// TIA Portal project "CHM_BORDEIRA_20190721" (V15) (continued)
REGION Network 14: I1.5 - CSW Valve Closed (CV-311)
   // True = CLOSED, False = NOT
   RUNG wire#powerrail
      Contact( "CSW Valve Closed" )
      I_Contact( "CSW Valve Open" )
      Coil( "10_DI_Data".CV311_CLSD )
   END_RUNG
   // the same network as SCL:
   "10_DI_Data".CV311_CLSD := "CSW Valve Closed" AND NOT "CSW Valve Open";
END_REGION

REGION Network 15: I1.6 - Flue Gas Scrubber CSW Valve Open (CV-312)
   // True = OPEN, False = NOT
   RUNG wire#powerrail
      Contact( "Flue Gas Scrubber CSW Valve Opened" )
      I_Contact( "Flue Gas Scrubber CSW Valve Closed" )
      Coil( "10_DI_Data".CV312_OPN )
   END_RUNG
   // the same network as SCL:
   "10_DI_Data".CV312_OPN := "Flue Gas Scrubber CSW Valve Opened" AND NOT "Flue Gas Scrubber CSW Valve Closed";
END_REGION

REGION Network 16: I1.7 - Flue Gas Scrubber CSW Valve Closed (CV-312)
   // True = CLOSED, False = NOT
   RUNG wire#powerrail
      Contact( "Flue Gas Scrubber CSW Valve Closed" )
      I_Contact( "Flue Gas Scrubber CSW Valve Opened" )
      Coil( "10_DI_Data".CV312_CLSD )
   END_RUNG
   // the same network as SCL:
   "10_DI_Data".CV312_CLSD := "Flue Gas Scrubber CSW Valve Closed" AND NOT "Flue Gas Scrubber CSW Valve Opened";
END_REGION

REGION Network 17: I2.0 - BC PLC Power Healthy
   // True = OK, False = NOK
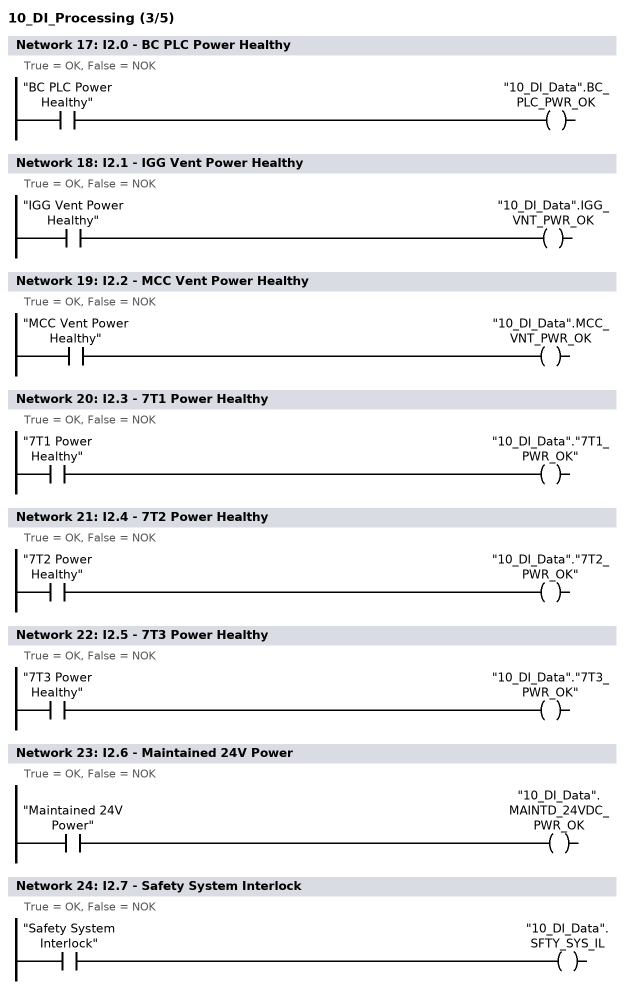
   RUNG wire#powerrail
      Contact( "BC PLC Power Healthy" )
      Coil( "10_DI_Data".BC_PLC_PWR_OK )
   END_RUNG
   // the same network as SCL:
   "10_DI_Data".BC_PLC_PWR_OK := "BC PLC Power Healthy";
END_REGION

REGION Network 18: I2.1 - IGG Vent Power Healthy
   // True = OK, False = NOK
   RUNG wire#powerrail
      Contact( "IGG Vent Power Healthy" )
      Coil( "10_DI_Data".IGG_VNT_PWR_OK )
   END_RUNG
   // the same network as SCL:
   "10_DI_Data".IGG_VNT_PWR_OK := "IGG Vent Power Healthy";
END_REGION

REGION Network 19: I2.2 - MCC Vent Power Healthy
   // True = OK, False = NOK
   RUNG wire#powerrail
      Contact( "MCC Vent Power Healthy" )
      Coil( "10_DI_Data".MCC_VNT_PWR_OK )
   END_RUNG
   // the same network as SCL:
   "10_DI_Data".MCC_VNT_PWR_OK := "MCC Vent Power Healthy";
END_REGION

REGION Network 20: I2.3 - 7T1 Power Healthy
   // True = OK, False = NOK
   RUNG wire#powerrail
      Contact( "7T1 Power Healthy" )
      Coil( "10_DI_Data"."7T1_PWR_OK" )
   END_RUNG
   // the same network as SCL:
   "10_DI_Data"."7T1_PWR_OK" := "7T1 Power Healthy";
END_REGION

REGION Network 21: I2.4 - 7T2 Power Healthy
   // True = OK, False = NOK
   RUNG wire#powerrail
      Contact( "7T2 Power Healthy" )
      Coil( "10_DI_Data"."7T2_PWR_OK" )
   END_RUNG
   // the same network as SCL:
   "10_DI_Data"."7T2_PWR_OK" := "7T2 Power Healthy";
END_REGION

REGION Network 22: I2.5 - 7T3 Power Healthy
   // True = OK, False = NOK
   RUNG wire#powerrail
      Contact( "7T3 Power Healthy" )
      Coil( "10_DI_Data"."7T3_PWR_OK" )
   END_RUNG
   // the same network as SCL:
   "10_DI_Data"."7T3_PWR_OK" := "7T3 Power Healthy";
END_REGION

REGION Network 23: I2.6 - Maintained 24V Power
   // True = OK, False = NOK
   RUNG wire#powerrail
      Contact( "Maintained 24V Power" )
      Coil( "10_DI_Data".MAINTD_24VDC_PWR_OK )
   END_RUNG
   // the same network as SCL:
   "10_DI_Data".MAINTD_24VDC_PWR_OK := "Maintained 24V Power";
END_REGION

REGION Network 24: I2.7 - Safety System Interlock
   // True = OK, False = NOK
   RUNG wire#powerrail
      Contact( "Safety System Interlock" )
      Coil( "10_DI_Data".SFTY_SYS_IL )
   END_RUNG
   // the same network as SCL:
   "10_DI_Data".SFTY_SYS_IL := "Safety System Interlock";
END_REGION

REGION Network 25: I3.0 - Cargo Blanketing IG Supply Valve Open (CV-432)
   // True = OPEN, False = NOT
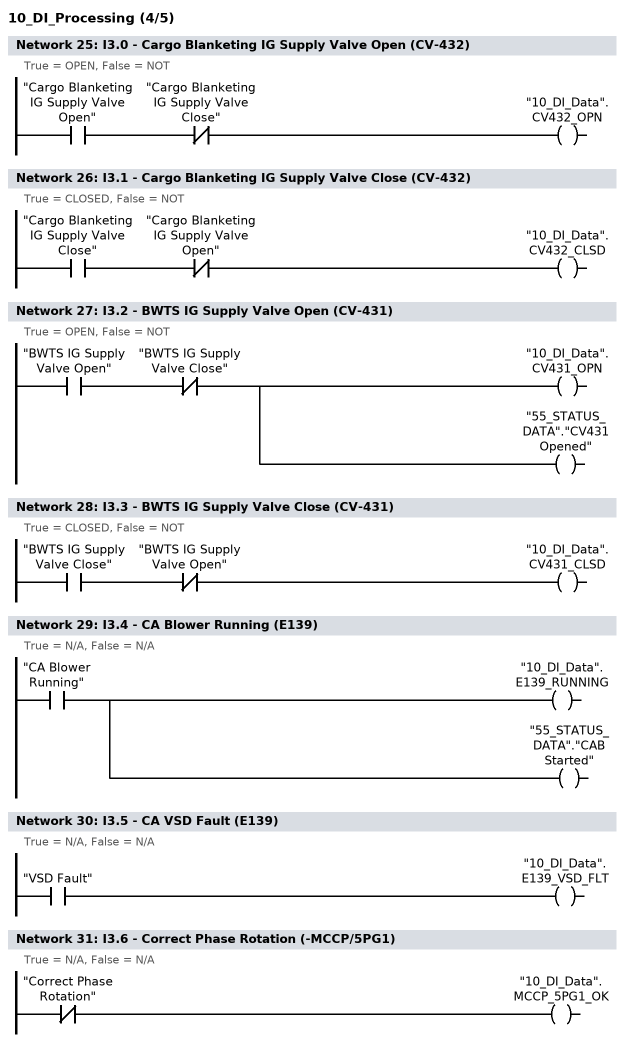
   RUNG wire#powerrail
      Contact( "Cargo Blanketing IG Supply Valve Open" )
      I_Contact( "Cargo Blanketing IG Supply Valve Close" )
      Coil( "10_DI_Data".CV432_OPN )
   END_RUNG
   // the same network as SCL:
   "10_DI_Data".CV432_OPN := "Cargo Blanketing IG Supply Valve Open" AND NOT "Cargo Blanketing IG Supply Valve Close";
END_REGION

REGION Network 26: I3.1 - Cargo Blanketing IG Supply Valve Close (CV-432)
   // True = CLOSED, False = NOT
   RUNG wire#powerrail
      Contact( "Cargo Blanketing IG Supply Valve Close" )
      I_Contact( "Cargo Blanketing IG Supply Valve Open" )
      Coil( "10_DI_Data".CV432_CLSD )
   END_RUNG
   // the same network as SCL:
   "10_DI_Data".CV432_CLSD := "Cargo Blanketing IG Supply Valve Close" AND NOT "Cargo Blanketing IG Supply Valve Open";
END_REGION

REGION Network 27: I3.2 - BWTS IG Supply Valve Open (CV-431)
   // True = OPEN, False = NOT
   RUNG wire#powerrail
      Contact( "BWTS IG Supply Valve Open" )
      I_Contact( "BWTS IG Supply Valve Close" )
      wire#w1
      Coil( "10_DI_Data".CV431_OPN )
   END_RUNG
   RUNG wire#w1
      Coil( "55_STATUS_DATA"."CV431 Opened" )
   END_RUNG
   // the same network as SCL:
   "10_DI_Data".CV431_OPN := "BWTS IG Supply Valve Open" AND NOT "BWTS IG Supply Valve Close";
   "55_STATUS_DATA"."CV431 Opened" := "10_DI_Data".CV431_OPN;
END_REGION

REGION Network 28: I3.3 - BWTS IG Supply Valve Close (CV-431)
   // True = CLOSED, False = NOT
   RUNG wire#powerrail
      Contact( "BWTS IG Supply Valve Close" )
      I_Contact( "BWTS IG Supply Valve Open" )
      Coil( "10_DI_Data".CV431_CLSD )
   END_RUNG
   // the same network as SCL:
   "10_DI_Data".CV431_CLSD := "BWTS IG Supply Valve Close" AND NOT "BWTS IG Supply Valve Open";
END_REGION

REGION Network 29: I3.4 - CA Blower Running (E139)
   // True = N/A, False = N/A
   RUNG wire#powerrail
      Contact( "CA Blower Running" )
      wire#w1
      Coil( "10_DI_Data".E139_RUNNING )
   END_RUNG
   RUNG wire#w1
      Coil( "55_STATUS_DATA"."CAB Started" )
   END_RUNG
   // the same network as SCL:
   "10_DI_Data".E139_RUNNING := "CA Blower Running";
   "55_STATUS_DATA"."CAB Started" := "CA Blower Running";
END_REGION

REGION Network 30: I3.5 - CA VSD Fault (E139)
   // True = N/A, False = N/A
   RUNG wire#powerrail
      Contact( "VSD Fault" )
      Coil( "10_DI_Data".E139_VSD_FLT )
   END_RUNG
   // the same network as SCL:
   "10_DI_Data".E139_VSD_FLT := "VSD Fault";
END_REGION

REGION Network 31: I3.6 - Correct Phase Rotation (-MCCP/5PG1)
   // True = N/A, False = N/A
   RUNG wire#powerrail
      I_Contact( "Correct Phase Rotation" )
      Coil( "10_DI_Data".MCCP_5PG1_OK )
   END_RUNG
   // the same network as SCL:
   "10_DI_Data".MCCP_5PG1_OK := NOT "Correct Phase Rotation";
END_REGION

REGION Network 32: I3.7 - Spare Input
   // True = N/A, False = N/A
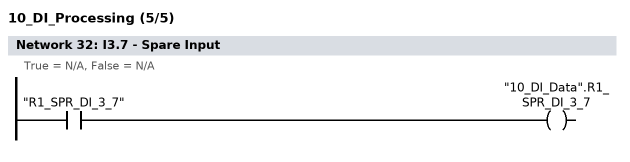
   RUNG wire#powerrail
      Contact( "R1_SPR_DI_3_7" )
      Coil( "10_DI_Data".R1_SPR_DI_3_7 )
   END_RUNG
   // the same network as SCL:
   "10_DI_Data".R1_SPR_DI_3_7 := "R1_SPR_DI_3_7";
END_REGION
END_FUNCTION

FUNCTION "12_AI_Processing" : Void   // FC12, LAD
TITLE = Analogue Input Processing
{ S7_Optimized_Access := 'TRUE' }
AUTHOR : JRS
VERSION : 0.1
// To process raw inputs prior to code use
BEGIN

REGION Network 1: IW112 - Combustion Air Pressure (PIT-102)
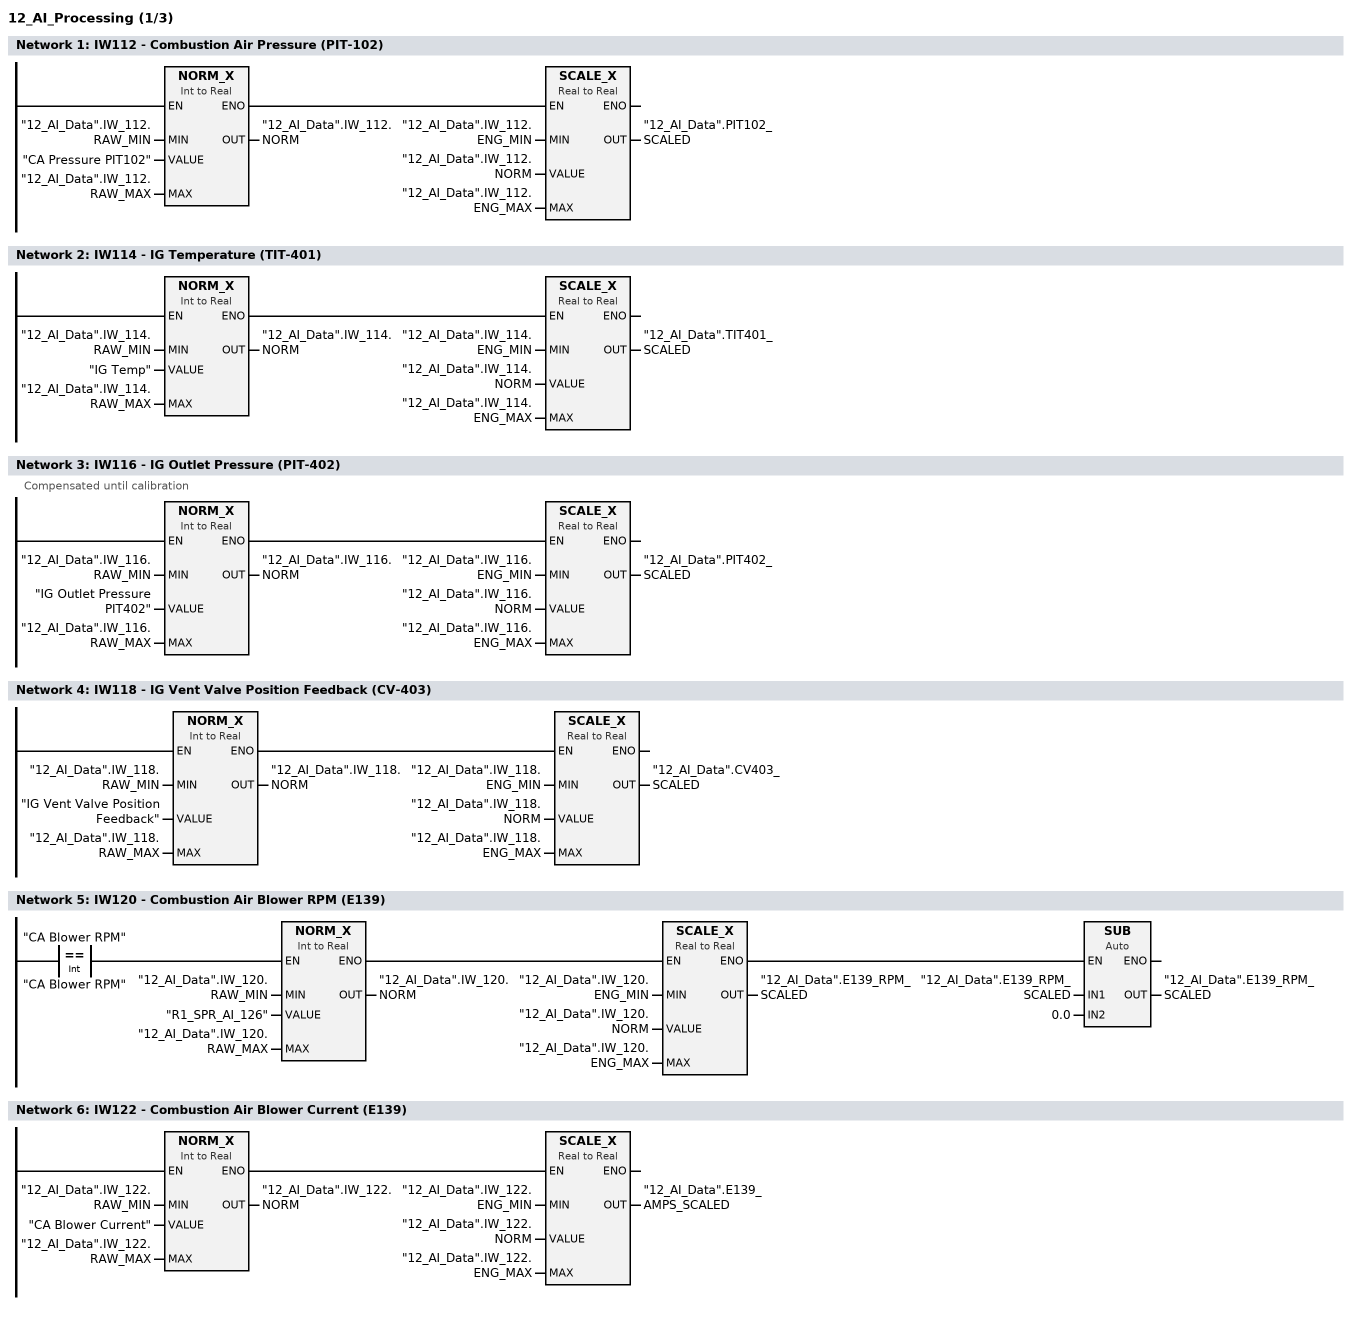
   RUNG wire#powerrail
      { S7_Templates := "[SrcType := Int, DestType := Real]" } Normalize(min := "12_AI_Data".IW_112.RAW_MIN, value := "CA Pressure PIT102", max := "12_AI_Data".IW_112.RAW_MAX, out => "12_AI_Data".IW_112.NORM)
      { S7_Templates := "[SrcType := Real, DestType := Real]" } Scale(min := "12_AI_Data".IW_112.ENG_MIN, value := "12_AI_Data".IW_112.NORM, max := "12_AI_Data".IW_112.ENG_MAX, out => "12_AI_Data".PIT102_SCALED)
   END_RUNG
   // the same network as SCL:
   "12_AI_Data".IW_112.NORM := NORM_X(MIN := "12_AI_Data".IW_112.RAW_MIN, VALUE := "CA Pressure PIT102", MAX := "12_AI_Data".IW_112.RAW_MAX);
   "12_AI_Data".PIT102_SCALED := SCALE_X(MIN := "12_AI_Data".IW_112.ENG_MIN, VALUE := "12_AI_Data".IW_112.NORM, MAX := "12_AI_Data".IW_112.ENG_MAX);
END_REGION

REGION Network 2: IW114 - IG Temperature (TIT-401)
   RUNG wire#powerrail
      { S7_Templates := "[SrcType := Int, DestType := Real]" } Normalize(min := "12_AI_Data".IW_114.RAW_MIN, value := "IG Temp", max := "12_AI_Data".IW_114.RAW_MAX, out => "12_AI_Data".IW_114.NORM)
      { S7_Templates := "[SrcType := Real, DestType := Real]" } Scale(min := "12_AI_Data".IW_114.ENG_MIN, value := "12_AI_Data".IW_114.NORM, max := "12_AI_Data".IW_114.ENG_MAX, out => "12_AI_Data".TIT401_SCALED)
   END_RUNG
   // the same network as SCL:
   "12_AI_Data".IW_114.NORM := NORM_X(MIN := "12_AI_Data".IW_114.RAW_MIN, VALUE := "IG Temp", MAX := "12_AI_Data".IW_114.RAW_MAX);
   "12_AI_Data".TIT401_SCALED := SCALE_X(MIN := "12_AI_Data".IW_114.ENG_MIN, VALUE := "12_AI_Data".IW_114.NORM, MAX := "12_AI_Data".IW_114.ENG_MAX);
END_REGION

REGION Network 3: IW116 - IG Outlet Pressure (PIT-402)
   // Compensated until calibration
   RUNG wire#powerrail
      { S7_Templates := "[SrcType := Int, DestType := Real]" } Normalize(min := "12_AI_Data".IW_116.RAW_MIN, value := "IG Outlet Pressure PIT402", max := "12_AI_Data".IW_116.RAW_MAX, out => "12_AI_Data".IW_116.NORM)
      { S7_Templates := "[SrcType := Real, DestType := Real]" } Scale(min := "12_AI_Data".IW_116.ENG_MIN, value := "12_AI_Data".IW_116.NORM, max := "12_AI_Data".IW_116.ENG_MAX, out => "12_AI_Data".PIT402_SCALED)
   END_RUNG
   // the same network as SCL:
   "12_AI_Data".IW_116.NORM := NORM_X(MIN := "12_AI_Data".IW_116.RAW_MIN, VALUE := "IG Outlet Pressure PIT402", MAX := "12_AI_Data".IW_116.RAW_MAX);
   "12_AI_Data".PIT402_SCALED := SCALE_X(MIN := "12_AI_Data".IW_116.ENG_MIN, VALUE := "12_AI_Data".IW_116.NORM, MAX := "12_AI_Data".IW_116.ENG_MAX);
END_REGION

REGION Network 4: IW118 - IG Vent Valve Position Feedback (CV-403)
   RUNG wire#powerrail
      { S7_Templates := "[SrcType := Int, DestType := Real]" } Normalize(min := "12_AI_Data".IW_118.RAW_MIN, value := "IG Vent Valve Position Feedback", max := "12_AI_Data".IW_118.RAW_MAX, out => "12_AI_Data".IW_118.NORM)
      { S7_Templates := "[SrcType := Real, DestType := Real]" } Scale(min := "12_AI_Data".IW_118.ENG_MIN, value := "12_AI_Data".IW_118.NORM, max := "12_AI_Data".IW_118.ENG_MAX, out => "12_AI_Data".CV403_SCALED)
   END_RUNG
   // the same network as SCL:
   "12_AI_Data".IW_118.NORM := NORM_X(MIN := "12_AI_Data".IW_118.RAW_MIN, VALUE := "IG Vent Valve Position Feedback", MAX := "12_AI_Data".IW_118.RAW_MAX);
   "12_AI_Data".CV403_SCALED := SCALE_X(MIN := "12_AI_Data".IW_118.ENG_MIN, VALUE := "12_AI_Data".IW_118.NORM, MAX := "12_AI_Data".IW_118.ENG_MAX);
END_REGION

REGION Network 5: IW120 - Combustion Air Blower RPM (E139)
   RUNG wire#powerrail
      { S7_Templates := "SrcType := Int" } EQ_Contact(in1 := "CA Blower RPM", in2 := "CA Blower RPM")
      { S7_Templates := "[SrcType := Int, DestType := Real]" } Normalize(min := "12_AI_Data".IW_120.RAW_MIN, value := "R1_SPR_AI_126", max := "12_AI_Data".IW_120.RAW_MAX, out => "12_AI_Data".IW_120.NORM)
      { S7_Templates := "[SrcType := Real, DestType := Real]" } Scale(min := "12_AI_Data".IW_120.ENG_MIN, value := "12_AI_Data".IW_120.NORM, max := "12_AI_Data".IW_120.ENG_MAX, out => "12_AI_Data".E139_RPM_SCALED)
      Sub(in1 := "12_AI_Data".E139_RPM_SCALED, in2 := 0.0, out => "12_AI_Data".E139_RPM_SCALED)
   END_RUNG
   // the same network as SCL:
   IF "CA Blower RPM" = "CA Blower RPM" THEN
       "12_AI_Data".IW_120.NORM := NORM_X(MIN := "12_AI_Data".IW_120.RAW_MIN, VALUE := "R1_SPR_AI_126", MAX := "12_AI_Data".IW_120.RAW_MAX);
       "12_AI_Data".E139_RPM_SCALED := SCALE_X(MIN := "12_AI_Data".IW_120.ENG_MIN, VALUE := "12_AI_Data".IW_120.NORM, MAX := "12_AI_Data".IW_120.ENG_MAX);
       "12_AI_Data".E139_RPM_SCALED := "12_AI_Data".E139_RPM_SCALED - 0.0;
   END_IF;
END_REGION

REGION Network 6: IW122 - Combustion Air Blower Current (E139)
   RUNG wire#powerrail
      { S7_Templates := "[SrcType := Int, DestType := Real]" } Normalize(min := "12_AI_Data".IW_122.RAW_MIN, value := "CA Blower Current", max := "12_AI_Data".IW_122.RAW_MAX, out => "12_AI_Data".IW_122.NORM)
      { S7_Templates := "[SrcType := Real, DestType := Real]" } Scale(min := "12_AI_Data".IW_122.ENG_MIN, value := "12_AI_Data".IW_122.NORM, max := "12_AI_Data".IW_122.ENG_MAX, out => "12_AI_Data".E139_AMPS_SCALED)
   END_RUNG
   // the same network as SCL:
   "12_AI_Data".IW_122.NORM := NORM_X(MIN := "12_AI_Data".IW_122.RAW_MIN, VALUE := "CA Blower Current", MAX := "12_AI_Data".IW_122.RAW_MAX);
   "12_AI_Data".E139_AMPS_SCALED := SCALE_X(MIN := "12_AI_Data".IW_122.ENG_MIN, VALUE := "12_AI_Data".IW_122.NORM, MAX := "12_AI_Data".IW_122.ENG_MAX);
END_REGION

REGION Network 7: IW124 - Fresh Water Bulk Tank Level (LIT-305)
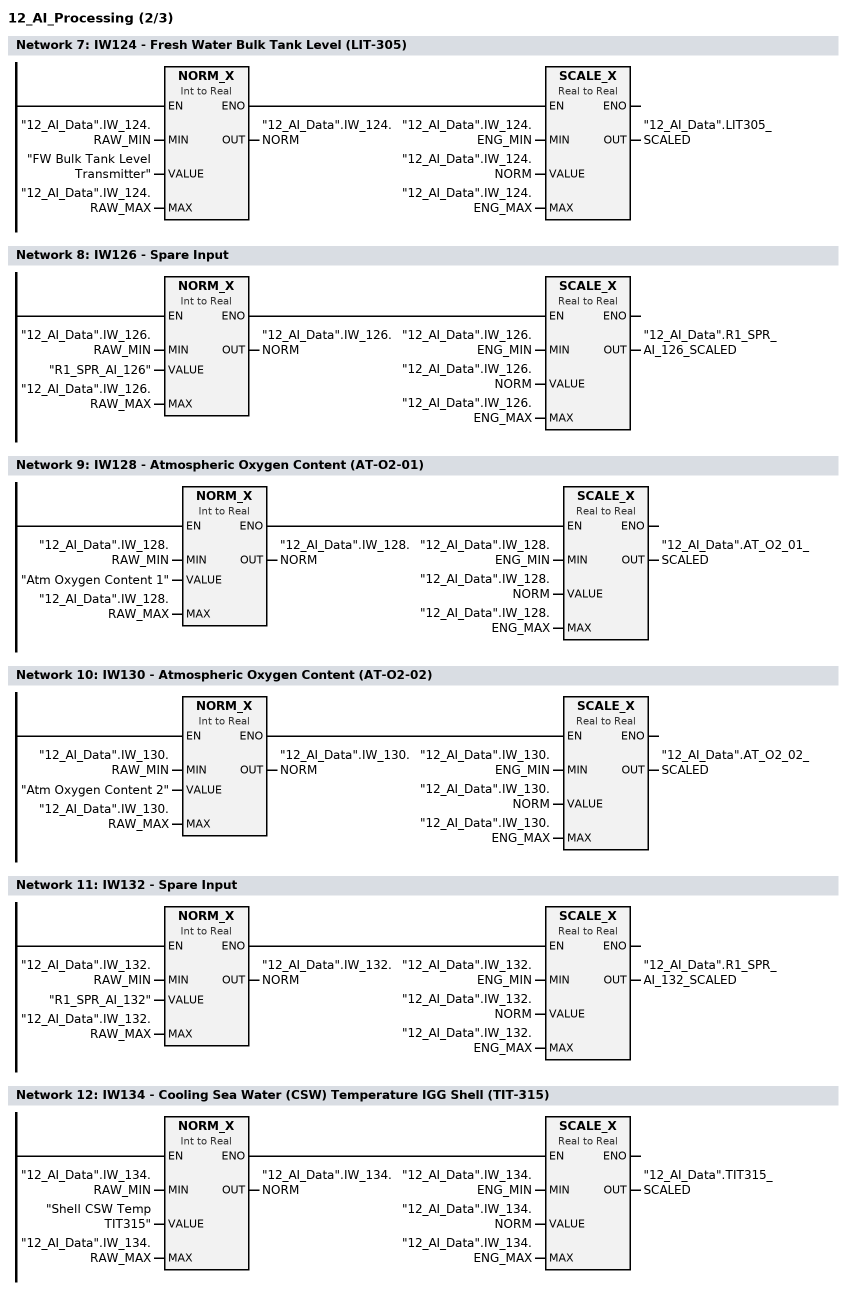
   RUNG wire#powerrail
      { S7_Templates := "[SrcType := Int, DestType := Real]" } Normalize(min := "12_AI_Data".IW_124.RAW_MIN, value := "FW Bulk Tank Level Transmitter", max := "12_AI_Data".IW_124.RAW_MAX, out => "12_AI_Data".IW_124.NORM)
      { S7_Templates := "[SrcType := Real, DestType := Real]" } Scale(min := "12_AI_Data".IW_124.ENG_MIN, value := "12_AI_Data".IW_124.NORM, max := "12_AI_Data".IW_124.ENG_MAX, out => "12_AI_Data".LIT305_SCALED)
   END_RUNG
   // the same network as SCL:
   "12_AI_Data".IW_124.NORM := NORM_X(MIN := "12_AI_Data".IW_124.RAW_MIN, VALUE := "FW Bulk Tank Level Transmitter", MAX := "12_AI_Data".IW_124.RAW_MAX);
   "12_AI_Data".LIT305_SCALED := SCALE_X(MIN := "12_AI_Data".IW_124.ENG_MIN, VALUE := "12_AI_Data".IW_124.NORM, MAX := "12_AI_Data".IW_124.ENG_MAX);
END_REGION

REGION Network 8: IW126 - Spare Input
   RUNG wire#powerrail
      { S7_Templates := "[SrcType := Int, DestType := Real]" } Normalize(min := "12_AI_Data".IW_126.RAW_MIN, value := "R1_SPR_AI_126", max := "12_AI_Data".IW_126.RAW_MAX, out => "12_AI_Data".IW_126.NORM)
      { S7_Templates := "[SrcType := Real, DestType := Real]" } Scale(min := "12_AI_Data".IW_126.ENG_MIN, value := "12_AI_Data".IW_126.NORM, max := "12_AI_Data".IW_126.ENG_MAX, out => "12_AI_Data".R1_SPR_AI_126_SCALED)
   END_RUNG
   // the same network as SCL:
   "12_AI_Data".IW_126.NORM := NORM_X(MIN := "12_AI_Data".IW_126.RAW_MIN, VALUE := "R1_SPR_AI_126", MAX := "12_AI_Data".IW_126.RAW_MAX);
   "12_AI_Data".R1_SPR_AI_126_SCALED := SCALE_X(MIN := "12_AI_Data".IW_126.ENG_MIN, VALUE := "12_AI_Data".IW_126.NORM, MAX := "12_AI_Data".IW_126.ENG_MAX);
END_REGION

REGION Network 9: IW128 - Atmospheric Oxygen Content (AT-O2-01)
   RUNG wire#powerrail
      { S7_Templates := "[SrcType := Int, DestType := Real]" } Normalize(min := "12_AI_Data".IW_128.RAW_MIN, value := "Atm Oxygen Content 1", max := "12_AI_Data".IW_128.RAW_MAX, out => "12_AI_Data".IW_128.NORM)
      { S7_Templates := "[SrcType := Real, DestType := Real]" } Scale(min := "12_AI_Data".IW_128.ENG_MIN, value := "12_AI_Data".IW_128.NORM, max := "12_AI_Data".IW_128.ENG_MAX, out => "12_AI_Data".AT_O2_01_SCALED)
   END_RUNG
   // the same network as SCL:
   "12_AI_Data".IW_128.NORM := NORM_X(MIN := "12_AI_Data".IW_128.RAW_MIN, VALUE := "Atm Oxygen Content 1", MAX := "12_AI_Data".IW_128.RAW_MAX);
   "12_AI_Data".AT_O2_01_SCALED := SCALE_X(MIN := "12_AI_Data".IW_128.ENG_MIN, VALUE := "12_AI_Data".IW_128.NORM, MAX := "12_AI_Data".IW_128.ENG_MAX);
END_REGION

REGION Network 10: IW130 - Atmospheric Oxygen Content (AT-O2-02)
   RUNG wire#powerrail
      { S7_Templates := "[SrcType := Int, DestType := Real]" } Normalize(min := "12_AI_Data".IW_130.RAW_MIN, value := "Atm Oxygen Content 2", max := "12_AI_Data".IW_130.RAW_MAX, out => "12_AI_Data".IW_130.NORM)
      { S7_Templates := "[SrcType := Real, DestType := Real]" } Scale(min := "12_AI_Data".IW_130.ENG_MIN, value := "12_AI_Data".IW_130.NORM, max := "12_AI_Data".IW_130.ENG_MAX, out => "12_AI_Data".AT_O2_02_SCALED)
   END_RUNG
   // the same network as SCL:
   "12_AI_Data".IW_130.NORM := NORM_X(MIN := "12_AI_Data".IW_130.RAW_MIN, VALUE := "Atm Oxygen Content 2", MAX := "12_AI_Data".IW_130.RAW_MAX);
   "12_AI_Data".AT_O2_02_SCALED := SCALE_X(MIN := "12_AI_Data".IW_130.ENG_MIN, VALUE := "12_AI_Data".IW_130.NORM, MAX := "12_AI_Data".IW_130.ENG_MAX);
END_REGION

REGION Network 11: IW132 - Spare Input
   RUNG wire#powerrail
      { S7_Templates := "[SrcType := Int, DestType := Real]" } Normalize(min := "12_AI_Data".IW_132.RAW_MIN, value := "R1_SPR_AI_132", max := "12_AI_Data".IW_132.RAW_MAX, out => "12_AI_Data".IW_132.NORM)
      { S7_Templates := "[SrcType := Real, DestType := Real]" } Scale(min := "12_AI_Data".IW_132.ENG_MIN, value := "12_AI_Data".IW_132.NORM, max := "12_AI_Data".IW_132.ENG_MAX, out => "12_AI_Data".R1_SPR_AI_132_SCALED)
   END_RUNG
   // the same network as SCL:
   "12_AI_Data".IW_132.NORM := NORM_X(MIN := "12_AI_Data".IW_132.RAW_MIN, VALUE := "R1_SPR_AI_132", MAX := "12_AI_Data".IW_132.RAW_MAX);
   "12_AI_Data".R1_SPR_AI_132_SCALED := SCALE_X(MIN := "12_AI_Data".IW_132.ENG_MIN, VALUE := "12_AI_Data".IW_132.NORM, MAX := "12_AI_Data".IW_132.ENG_MAX);
END_REGION

REGION Network 12: IW134 - Cooling Sea Water (CSW) Temperature IGG Shell (TIT-315)
   RUNG wire#powerrail
      { S7_Templates := "[SrcType := Int, DestType := Real]" } Normalize(min := "12_AI_Data".IW_134.RAW_MIN, value := "Shell CSW Temp TIT315", max := "12_AI_Data".IW_134.RAW_MAX, out => "12_AI_Data".IW_134.NORM)
      { S7_Templates := "[SrcType := Real, DestType := Real]" } Scale(min := "12_AI_Data".IW_134.ENG_MIN, value := "12_AI_Data".IW_134.NORM, max := "12_AI_Data".IW_134.ENG_MAX, out => "12_AI_Data".TIT315_SCALED)
   END_RUNG
   // the same network as SCL:
   "12_AI_Data".IW_134.NORM := NORM_X(MIN := "12_AI_Data".IW_134.RAW_MIN, VALUE := "Shell CSW Temp TIT315", MAX := "12_AI_Data".IW_134.RAW_MAX);
   "12_AI_Data".TIT315_SCALED := SCALE_X(MIN := "12_AI_Data".IW_134.ENG_MIN, VALUE := "12_AI_Data".IW_134.NORM, MAX := "12_AI_Data".IW_134.ENG_MAX);
END_REGION

REGION Network 13: IW136 - Cooling Sea Water (CSW) Temperature IGG Inlet (TIT_319)
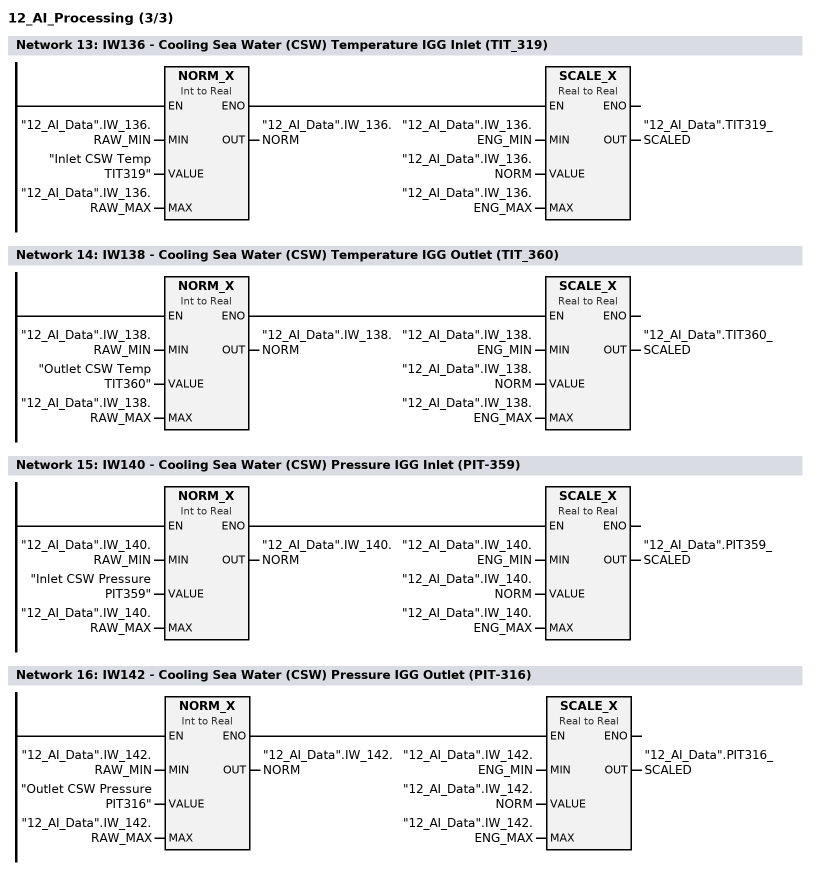
   RUNG wire#powerrail
      { S7_Templates := "[SrcType := Int, DestType := Real]" } Normalize(min := "12_AI_Data".IW_136.RAW_MIN, value := "Inlet CSW Temp TIT319", max := "12_AI_Data".IW_136.RAW_MAX, out => "12_AI_Data".IW_136.NORM)
      { S7_Templates := "[SrcType := Real, DestType := Real]" } Scale(min := "12_AI_Data".IW_136.ENG_MIN, value := "12_AI_Data".IW_136.NORM, max := "12_AI_Data".IW_136.ENG_MAX, out => "12_AI_Data".TIT319_SCALED)
   END_RUNG
   // the same network as SCL:
   "12_AI_Data".IW_136.NORM := NORM_X(MIN := "12_AI_Data".IW_136.RAW_MIN, VALUE := "Inlet CSW Temp TIT319", MAX := "12_AI_Data".IW_136.RAW_MAX);
   "12_AI_Data".TIT319_SCALED := SCALE_X(MIN := "12_AI_Data".IW_136.ENG_MIN, VALUE := "12_AI_Data".IW_136.NORM, MAX := "12_AI_Data".IW_136.ENG_MAX);
END_REGION

REGION Network 14: IW138 - Cooling Sea Water (CSW) Temperature IGG Outlet (TIT_360)
   RUNG wire#powerrail
      { S7_Templates := "[SrcType := Int, DestType := Real]" } Normalize(min := "12_AI_Data".IW_138.RAW_MIN, value := "Outlet CSW Temp TIT360", max := "12_AI_Data".IW_138.RAW_MAX, out => "12_AI_Data".IW_138.NORM)
      { S7_Templates := "[SrcType := Real, DestType := Real]" } Scale(min := "12_AI_Data".IW_138.ENG_MIN, value := "12_AI_Data".IW_138.NORM, max := "12_AI_Data".IW_138.ENG_MAX, out => "12_AI_Data".TIT360_SCALED)
   END_RUNG
   // the same network as SCL:
   "12_AI_Data".IW_138.NORM := NORM_X(MIN := "12_AI_Data".IW_138.RAW_MIN, VALUE := "Outlet CSW Temp TIT360", MAX := "12_AI_Data".IW_138.RAW_MAX);
   "12_AI_Data".TIT360_SCALED := SCALE_X(MIN := "12_AI_Data".IW_138.ENG_MIN, VALUE := "12_AI_Data".IW_138.NORM, MAX := "12_AI_Data".IW_138.ENG_MAX);
END_REGION

REGION Network 15: IW140 - Cooling Sea Water (CSW) Pressure IGG Inlet (PIT-359)
   RUNG wire#powerrail
      { S7_Templates := "[SrcType := Int, DestType := Real]" } Normalize(min := "12_AI_Data".IW_140.RAW_MIN, value := "Inlet CSW Pressure PIT359", max := "12_AI_Data".IW_140.RAW_MAX, out => "12_AI_Data".IW_140.NORM)
      { S7_Templates := "[SrcType := Real, DestType := Real]" } Scale(min := "12_AI_Data".IW_140.ENG_MIN, value := "12_AI_Data".IW_140.NORM, max := "12_AI_Data".IW_140.ENG_MAX, out => "12_AI_Data".PIT359_SCALED)
   END_RUNG
   // the same network as SCL:
   "12_AI_Data".IW_140.NORM := NORM_X(MIN := "12_AI_Data".IW_140.RAW_MIN, VALUE := "Inlet CSW Pressure PIT359", MAX := "12_AI_Data".IW_140.RAW_MAX);
   "12_AI_Data".PIT359_SCALED := SCALE_X(MIN := "12_AI_Data".IW_140.ENG_MIN, VALUE := "12_AI_Data".IW_140.NORM, MAX := "12_AI_Data".IW_140.ENG_MAX);
END_REGION

REGION Network 16: IW142 - Cooling Sea Water (CSW) Pressure IGG Outlet (PIT-316)
   RUNG wire#powerrail
      { S7_Templates := "[SrcType := Int, DestType := Real]" } Normalize(min := "12_AI_Data".IW_142.RAW_MIN, value := "Outlet CSW Pressure PIT316", max := "12_AI_Data".IW_142.RAW_MAX, out => "12_AI_Data".IW_142.NORM)
      { S7_Templates := "[SrcType := Real, DestType := Real]" } Scale(min := "12_AI_Data".IW_142.ENG_MIN, value := "12_AI_Data".IW_142.NORM, max := "12_AI_Data".IW_142.ENG_MAX, out => "12_AI_Data".PIT316_SCALED)
   END_RUNG
   // the same network as SCL:
   "12_AI_Data".IW_142.NORM := NORM_X(MIN := "12_AI_Data".IW_142.RAW_MIN, VALUE := "Outlet CSW Pressure PIT316", MAX := "12_AI_Data".IW_142.RAW_MAX);
   "12_AI_Data".PIT316_SCALED := SCALE_X(MIN := "12_AI_Data".IW_142.ENG_MIN, VALUE := "12_AI_Data".IW_142.NORM, MAX := "12_AI_Data".IW_142.ENG_MAX);
END_REGION
END_FUNCTION

FUNCTION "14_DQ_Processing" : Void   // FC14, LAD
TITLE = Digital Output Processing
{ S7_Optimized_Access := 'TRUE' }
AUTHOR : JRS
VERSION : 0.1
// To process code outputs prior to physical connection
   VAR_TEMP
      RET_VAL_1 : Int;
   END_VAR
   VAR_TEMP   // added for the SCL form of the ladder/FBD networks
      _w1 : Bool;
      _w2 : Bool;
   END_VAR
BEGIN

REGION Network 1: Q0.0 - Fuel Pump #1 Control (E-500-A)
   // True = RUN, False = NOT
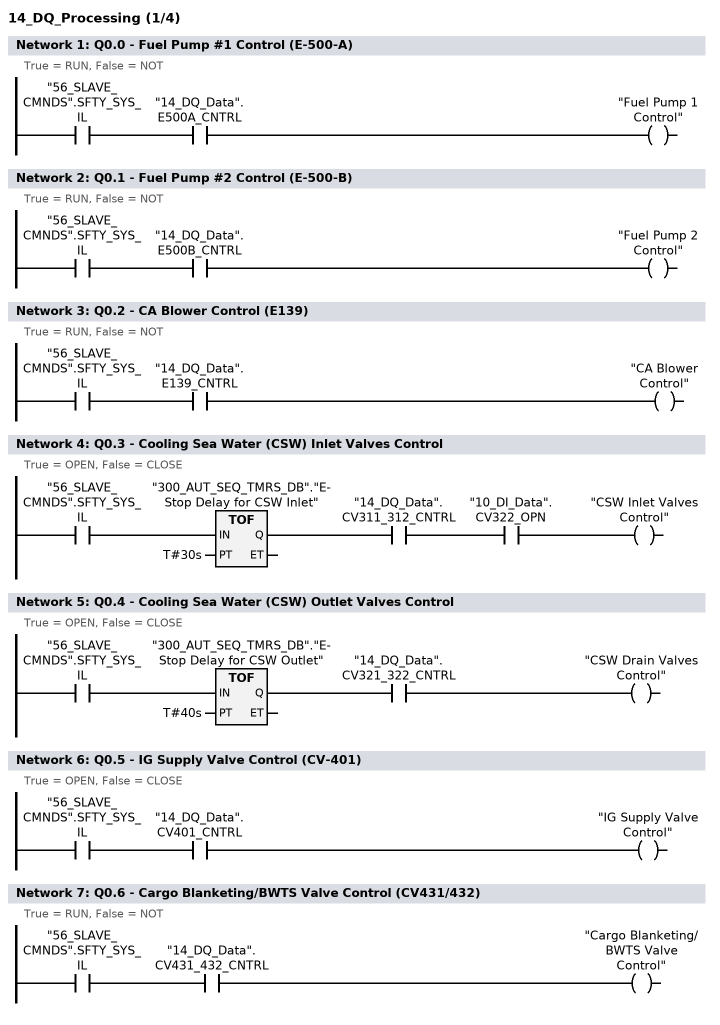
   RUNG wire#powerrail
      Contact( "56_SLAVE_CMNDS".SFTY_SYS_IL )
      Contact( "14_DQ_Data".E500A_CNTRL )
      Coil( "Fuel Pump 1 Control" )
   END_RUNG
   // the same network as SCL:
   "Fuel Pump 1 Control" := "56_SLAVE_CMNDS".SFTY_SYS_IL AND "14_DQ_Data".E500A_CNTRL;
END_REGION

REGION Network 2: Q0.1 - Fuel Pump #2 Control (E-500-B)
   // True = RUN, False = NOT
   RUNG wire#powerrail
      Contact( "56_SLAVE_CMNDS".SFTY_SYS_IL )
      Contact( "14_DQ_Data".E500B_CNTRL )
      Coil( "Fuel Pump 2 Control" )
   END_RUNG
   // the same network as SCL:
   "Fuel Pump 2 Control" := "56_SLAVE_CMNDS".SFTY_SYS_IL AND "14_DQ_Data".E500B_CNTRL;
END_REGION

REGION Network 3: Q0.2 - CA Blower Control (E139)
   // True = RUN, False = NOT
   RUNG wire#powerrail
      Contact( "56_SLAVE_CMNDS".SFTY_SYS_IL )
      Contact( "14_DQ_Data".E139_CNTRL )
      Coil( "CA Blower Control" )
   END_RUNG
   // the same network as SCL:
   "CA Blower Control" := "56_SLAVE_CMNDS".SFTY_SYS_IL AND "14_DQ_Data".E139_CNTRL;
END_REGION

REGION Network 4: Q0.3 - Cooling Sea Water (CSW) Inlet Valves Control
   // True = OPEN, False = CLOSE
   "300_AUT_SEQ_TMRS_DB"."E-Stop Delay for CSW Inlet".TOF(IN := "56_SLAVE_CMNDS".SFTY_SYS_IL, PT := T#30s);
   "CSW Inlet Valves Control" := "300_AUT_SEQ_TMRS_DB"."E-Stop Delay for CSW Inlet".Q AND "14_DQ_Data".CV311_312_CNTRL AND "10_DI_Data".CV322_OPN;
END_REGION

REGION Network 5: Q0.4 - Cooling Sea Water (CSW) Outlet Valves Control
   // True = OPEN, False = CLOSE
   "300_AUT_SEQ_TMRS_DB"."E-Stop Delay for CSW Outlet".TOF(IN := "56_SLAVE_CMNDS".SFTY_SYS_IL, PT := T#40s);
   "CSW Drain Valves Control" := "300_AUT_SEQ_TMRS_DB"."E-Stop Delay for CSW Outlet".Q AND "14_DQ_Data".CV321_322_CNTRL;
END_REGION

REGION Network 6: Q0.5 - IG Supply Valve Control (CV-401)
   // True = OPEN, False = CLOSE
   RUNG wire#powerrail
      Contact( "56_SLAVE_CMNDS".SFTY_SYS_IL )
      Contact( "14_DQ_Data".CV401_CNTRL )
      Coil( "IG Supply Valve Control" )
   END_RUNG
   // the same network as SCL:
   "IG Supply Valve Control" := "56_SLAVE_CMNDS".SFTY_SYS_IL AND "14_DQ_Data".CV401_CNTRL;
END_REGION

REGION Network 7: Q0.6 - Cargo Blanketing/BWTS Valve Control (CV431/432)
   // True = RUN, False = NOT
   RUNG wire#powerrail
      Contact( "56_SLAVE_CMNDS".SFTY_SYS_IL )
      Contact( "14_DQ_Data".CV431_432_CNTRL )
      Coil( "Cargo Blanketing/BWTS Valve Control" )
   END_RUNG
   // the same network as SCL:
   "Cargo Blanketing/BWTS Valve Control" := "56_SLAVE_CMNDS".SFTY_SYS_IL AND "14_DQ_Data".CV431_432_CNTRL;
END_REGION

REGION Network 8: Q0.7 - Spare Output
   // True = RUN, False = NOT
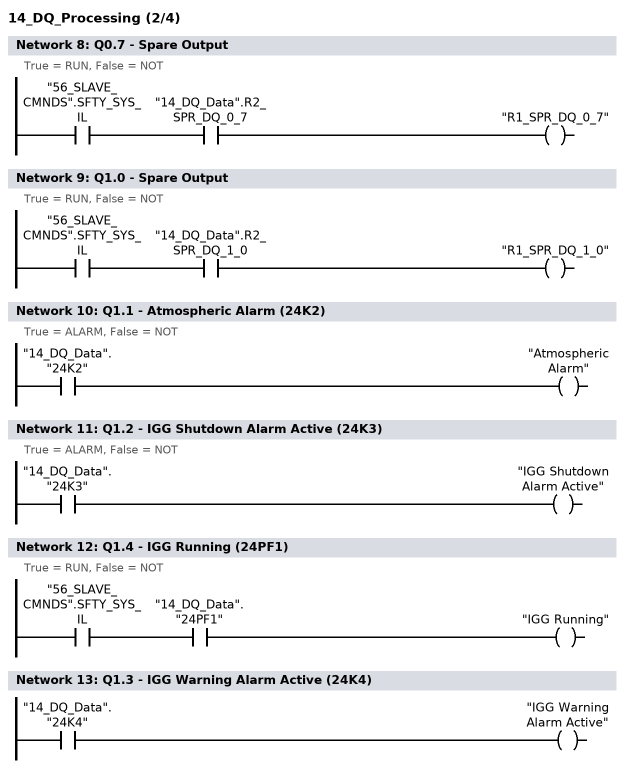
   RUNG wire#powerrail
      Contact( "56_SLAVE_CMNDS".SFTY_SYS_IL )
      Contact( "14_DQ_Data".R2_SPR_DQ_0_7 )
      Coil( "R1_SPR_DQ_0_7" )
   END_RUNG
   // the same network as SCL:
   "R1_SPR_DQ_0_7" := "56_SLAVE_CMNDS".SFTY_SYS_IL AND "14_DQ_Data".R2_SPR_DQ_0_7;
END_REGION

REGION Network 9: Q1.0 - Spare Output
   // True = RUN, False = NOT
   RUNG wire#powerrail
      Contact( "56_SLAVE_CMNDS".SFTY_SYS_IL )
      Contact( "14_DQ_Data".R2_SPR_DQ_1_0 )
      Coil( "R1_SPR_DQ_1_0" )
   END_RUNG
   // the same network as SCL:
   "R1_SPR_DQ_1_0" := "56_SLAVE_CMNDS".SFTY_SYS_IL AND "14_DQ_Data".R2_SPR_DQ_1_0;
END_REGION

REGION Network 10: Q1.1 - Atmospheric Alarm (24K2)
   // True = ALARM, False = NOT
   RUNG wire#powerrail
      Contact( "14_DQ_Data"."24K2" )
      Coil( "Atmospheric Alarm" )
   END_RUNG
   // the same network as SCL:
   "Atmospheric Alarm" := "14_DQ_Data"."24K2";
END_REGION

REGION Network 11: Q1.2 - IGG Shutdown Alarm Active (24K3)
   // True = ALARM, False = NOT
   RUNG wire#powerrail
      Contact( "14_DQ_Data"."24K3" )
      Coil( "IGG Shutdown Alarm Active" )
   END_RUNG
   // the same network as SCL:
   "IGG Shutdown Alarm Active" := "14_DQ_Data"."24K3";
END_REGION

REGION Network 12: Q1.4 - IGG Running (24PF1)
   // True = RUN, False = NOT
   RUNG wire#powerrail
      Contact( "56_SLAVE_CMNDS".SFTY_SYS_IL )
      Contact( "14_DQ_Data"."24PF1" )
      Coil( "IGG Running" )
   END_RUNG
   // the same network as SCL:
   "IGG Running" := "56_SLAVE_CMNDS".SFTY_SYS_IL AND "14_DQ_Data"."24PF1";
END_REGION

REGION Network 13: Q1.3 - IGG Warning Alarm Active (24K4)
   RUNG wire#powerrail
      Contact( "14_DQ_Data"."24K4" )
      Coil( "IGG Warning Alarm Active" )
   END_RUNG
   // the same network as SCL:
   "IGG Warning Alarm Active" := "14_DQ_Data"."24K4";
END_REGION

